
       // Clear the Array and start the request
       IF #wSDOStatus = 12 THEN //Step 12
           FILL_BLK(IN := 0,
                    COUNT := 64,
                    OUT => #bySDODataArray[0]);
           #bSDOReq := TRUE;
           #bSDOWriteDone := FALSE;
           #wSDOStatus := 13; //proceed to Step 13
       END_IF;
       // setup the array data and start WRREC
       IF #wSDOStatus = 13 THEN //Step 13
           #bySDODataArray[0] := 16#f9; //Request Reference
           #bySDODataArray[1] := 16#02; //2 for write PNU
           #bySDODataArray[2] := 16#00; //Axis# is 0 for AKD
           #bySDODataArray[3] := 16#01; // Number of parameters to write at a time
           // Set PNU 916 subindex 5
           #bySDODataArray[4] := 16#10; //Attribute is 0x10
           #bySDODataArray[5] := 16#01; //Number of elements =1
           #bySDODataArray[6] := 16#03; //0x394 for PNU 916
           #bySDODataArray[7] := 16#94; //PNU 916
           #bySDODataArray[8] := 16#00; //subindex
           #bySDODataArray[9] := 16#05; //subindex 5 for 6th word of telegram
           // To PNU 52 (ITIST_GLATT)
           #bySDODataArray[10] := 16#42; //Format =0x42 for Word
           #bySDODataArray[11] := 16#01; //Number of values
           #bySDODataArray[12] := 16#00; //data
           #bySDODataArray[13] := 16#34; //data - Signal #52 (0x34) for ITIST_GLATT (IL.FB)

           #SDOWrite(REQ := #bSDOReq, //do the PNU write
                     ID := #iID,
                     INDEX := 47, //AKD suppors "Record Data 47"
                     LEN := 14,   //data length
                     BUSY => #bSDOWriteBusy,
                     DONE => #bSDOWriteDone,
                     ERROR => #bSDOWriteError,
                     RECORD := #bySDODataArray);
           IF #bSDOWriteBusy THEN
               #bSDOReq := FALSE;
           ELSIF #bSDOWriteDone THEN
               #wSDOStatus := 14; //proceed to Step 14
               //#oInitDone := 1;    //telegram configuration complete
           END_IF;
       END_IF;

       // Set OpMode 
       // Clear the Array and start the request
       IF #wSDOStatus = 14 THEN //Step 14
           FILL_BLK(IN := 0,
                    COUNT := 64,
                    OUT => #bySDODataArray[0]);
           #bSDOReq := TRUE;
           #bSDOWriteDone := FALSE;
           #wSDOStatus := 15; //proceed to Step 15
       END_IF;
       // Set OpMode = 2 Position
       IF #wSDOStatus = 15 THEN //Step 15
           #bySDODataArray[0] := 16#fe; //Request Reference
           #bySDODataArray[1] := 16#02; //2 for write PNU
           #bySDODataArray[2] := 16#00; //Axis# is 0 for AKD
           #bySDODataArray[3] := 16#01; // Number of parameters to write at a time
               // Set PNU 930 subindex 0 (DRV.OPMODE)
           #bySDODataArray[4] := 16#10; //Attribute is 0x10
           #bySDODataArray[5] := 16#01; //Number of elements =1
           #bySDODataArray[6] := 16#03; //0x3A2 for PNU 930 - opmode
           #bySDODataArray[7] := 16#A2; //PNU 930
           #bySDODataArray[8] := 16#00; //subindex 0
           #bySDODataArray[9] := 16#00; //subindex 0
               // To 2 (position mode)
           #bySDODataArray[10] := 16#42; //Format =0x42 for Word
           #bySDODataArray[11] := 16#01; //Number of values
           #bySDODataArray[12] := 16#02; //data
           #bySDODataArray[13] := 16#02; //data - vlaue = 2 for position mode

           #SDOWrite(REQ := #bSDOReq, //do the PNU write
                     ID := #iID,
                     INDEX := 47, //AKD suppors "Record Data 47"
                     LEN := 14,   //data length
                     BUSY => #bSDOWriteBusy,
                     DONE => #bSDOWriteDone,
                     ERROR => #bSDOWriteError,
                     RECORD := #bySDODataArray);
           IF #bSDOWriteBusy THEN
               #bSDOReq := FALSE;
           ELSIF #bSDOWriteDone THEN
               #wSDOStatus := 20; // setup complete - skip to process
               #oInitDone := TRUE;    //telegram configuration complete
           END_IF;
       END_IF;
   END_IF;

   // Read ZSW and set output values
   IF NOT #iInit AND #wSDOStatus > 19 THEN
       #wPNReadStatus := DPRD_DAT(LADDR := #iID,
                                  RECORD => #TG_400.Receive);
       IF #wPNReadStatus = 0 THEN
           #bPNReadError := FALSE;

           #oStatus.%W0 := #TG_400.Receive.ZSW1;
           IF #wSDOStatus > 20 THEN
               #oStatus.%W1 := #wSDOReadValue;
           ELSE
               #oStatus.%W1 := 0;
           END_IF;
           #oPos.%W0 := #TG_400.Receive.XIST_A_1;
           #oPos.%W1 := #TG_400.Receive.XIST_A;
           #oVel := #TG_400.Receive.NIST_A;
           #oCurrent := #TG_400.Receive.ITIST_GLATT;

           #oEnabled := #TG_400.Receive.ZSW1.%X0 AND #TG_400.Receive.ZSW1.%X1 AND #TG_400.Receive.ZSW1.%X2 AND NOT #TG_400.Receive.ZSW1.%X6;
           #oFault := #TG_400.Receive.ZSW1.%X3;
           #oMoving := NOT #TG_400.Receive.ZSW1.%X13 OR #TG_400.Receive.ZSW1.%X14 OR #TG_400.Receive.ZSW1.%X12;
           #oHomed := #TG_400.Receive.ZSW1.%X11;
           IF #TG_400.Send.STW1.%X6 THEN        // Reset the InPos Flag for a minimum of one write cycle
               #oInPos := FALSE;
           ELSE
               #oInPos := #TG_400.Receive.ZSW1.%X10;
           END_IF;
           #oWarning := #TG_400.Receive.ZSW1.%X7;
       ELSE
           #bPNReadError := TRUE;
       END_IF;

   END_IF;

   // Do the write always as the zero Telegramm needs to be send on a init aswell
   #wPNWriteStatus := DPWR_DAT(LADDR := #iID,
                               RECORD := #TG_400.Send);

   // set STW1 and values for the AKD
   IF NOT #iInit AND #wSDOStatus > 19 THEN
       IF #wPNWriteStatus = 0 THEN
           #bPNWriteError := FALSE;

           #TG_400.Send.STW1.%X10 := TRUE;
           IF #TG_400.Receive.ZSW1.%X9 THEN     // PLC has control

               // Do a EStop
               IF #iEStop THEN
                   #TG_400.Send.STW1.%X2 := FALSE;
                   #bEstop := TRUE;
               END_IF;

               // Do a reset
               IF #iReset AND NOT #bResetDone THEN
                   #wSDOStatus := 20;
                   #TG_400.Send.STW1.%X7 := TRUE;
                   #bResetDone := TRUE;
                   #bEstop := FALSE;
                   #wStartReset := #TG_400.Receive.ZSW2;
               END_IF;
               IF ABS(#wStartReset - #TG_400.Receive.ZSW2) > 2 THEN
                   #TG_400.Send.STW1.%X7 := FALSE;
               END_IF;

               // Enable the drive
               IF #iSW_Enable AND NOT #bEstop AND NOT (#bSWEnabled AND #TG_400.Receive.ZSW1.%X6 OR #TG_400.Receive.ZSW1.%X3) THEN
                   IF #TG_400.Receive.ZSW1.%X6 THEN      // Switch on inhibited
                       #TG_400.Send.STW1.%X1 := TRUE;
                       #TG_400.Send.STW1.%X2 := TRUE;
                   ELSE
                       IF #TG_400.Receive.ZSW1.%X0 THEN     // Ready for switiching on
                           #TG_400.Send.STW1.%X0 := TRUE;
                           IF #TG_400.Receive.ZSW1.%X1 THEN       // Switched on
                               #TG_400.Send.STW1.%X3 := TRUE;
                               IF #TG_400.Receive.ZSW1.%X2 THEN       // Operation
                                   #TG_400.Send.STW1.%X12 := TRUE; //turn on real time jogging mode
                                   #bSWEnabled := TRUE;

                                   // Do a Stop
                                   IF #iStop THEN
                                       #TG_400.Send.STW1.%X4 := FALSE;   // Stop active motion task
                                       #TG_400.Send.STW1.%X5 := FALSE;   // Stop active motion task
                                       #TG_400.Send.STW1.%X8 := FALSE;   // Stop jog 1
                                       #TG_400.Send.STW1.%X9 := FALSE;   // Stop jog 2
                                       #TG_400.Send.STW1.%X11 := FALSE;  // Stop homeing
                                       //#TG_400.Send.STW1.%X12 := FALSE;  // Stop real time jogging mode
                                   ELSE

                                       // Do home
                                       IF #iStart_Homing AND NOT #bHomeStarted THEN
                                           #TG_400.Send.HOME_DIST := #iCmdPos.%W1;
                                           #TG_400.Send.HOME_DIST_1 := #iCmdPos.%W0;
                                           #TG_400.Send.STW1.%X11 := TRUE;
                                           #wHomingStartPoint := #TG_400.Receive.ZSW2;
                                           #bHomeStarted := TRUE;
                                       ELSE
                                           IF #TG_400.Receive.ZSW1.%X11 AND #TG_400.Receive.ZSW1.%X13 AND (ABS(#wHomingStartPoint - #TG_400.Receive.ZSW2) > 5) THEN
                                               #TG_400.Send.STW1.%X11 := FALSE;
                                           END_IF;

                                           // Jogging
                                           IF #iStart_Jog AND #iCmdVel <> 0 THEN
                                               #TG_400.Send.STW1.%X8 := TRUE;
                                               //#TG_400.Send.STW1.%X12 := TRUE;

                                               // if the speed input is negative set Bit 13 for reverse direction 
                                               IF #iCmdVel.%X31 = 1 THEN
                                                   #TG_400.Send.STW1.%X13 := TRUE;
                                                   #TG_400.Send.MDI_VELOCITY := (16#ffff - #iCmdVel.%W1 + 1);
                                                   #TG_400.Send.MDI_VELOCITY_1 := (16#ffff - #iCmdVel.%W0 + 1);
                                               ELSE
                                                   #TG_400.Send.STW1.%X13 := FALSE;
                                                   #TG_400.Send.MDI_VELOCITY := #iCmdVel.%W1;
                                                   #TG_400.Send.MDI_VELOCITY_1 := #iCmdVel.%W0;
                                               END_IF;

                                               #TG_400.Send.MDI_ACC := #iCmdAcc;
                                               #TG_400.Send.MDI_DEC := #iCmdDec;
                                           ELSE
                                               #TG_400.Send.STW1.%X8 := FALSE;
                                               //#TG_400.Send.STW1.%X12 := FALSE;

                                               // Interrupt a move
                                               IF #iMT_Pause THEN
                                                   #TG_400.Send.STW1.%X5 := FALSE;    // intermediate stop, motion is paused and will continue when the pause is lifted
                                               ELSE
                                                   #TG_400.Send.STW1.%X5 := TRUE;    // No intermediate stop
                                               END_IF;

                                               // Reset the rising edge of the start bit to be read for the next task
                                               IF #TG_400.Receive.ZSW1.%X12 OR ABS(#wStartMove - #TG_400.Receive.ZSW2) > 62 THEN //if start command has been acknowledged, or >62 telegram transmissions
                                                   #bStartMoveDone := TRUE; // the process to start the move has been completed
                                                   #TG_400.Send.STW1.%X6 := FALSE; //turn off the start bit
                                               END_IF;
                                               // Move
                                               IF #iStart_Move AND NOT #bStartMove THEN
                                                   #TG_400.Send.MDI_MOD := #iMT_MoveType;   // 1 = absolute, 0 = relative
                                                   #TG_400.Send.SATZANW := #iMTNum;      // 0x8000 = direct motion task, otherwise select a motion task from the AKD
                                                   #TG_400.Send.MDI_TARPOS := #iCmdPos.%W1;
                                                   #TG_400.Send.MDI_TARPOS_1 := #iCmdPos.%W0;
                                                   #TG_400.Send.MDI_VELOCITY := #iCmdVel.%W1;
                                                   #TG_400.Send.MDI_VELOCITY_1 := #iCmdVel.%W0;
                                                   #TG_400.Send.MDI_ACC := #iCmdAcc;
                                                   #TG_400.Send.MDI_DEC := #iCmdDec;
                                                   #TG_400.Send.STW1.%X4 := TRUE;    // Do not reject traversing task
                                                   #TG_400.Send.STW1.%X5 := TRUE;    // No intermediate stop
                                                   #TG_400.Send.STW1.%X6 := TRUE;    // Start the move

                                                   #bStartMove := TRUE; // the process to start the move has been started but not completed
                                                   #bStartMoveDone := FALSE; // the process to start the move has not been completed
                                                   #wStartMove := #TG_400.Receive.ZSW2;
                                               END_IF; //If Start move

                                           END_IF; //If Start Jog
                                       END_IF; //If Start Homing
                                   END_IF; // If Stop
                               END_IF; // If ZSW1 bit2 Operation Enabled
                           END_IF; // If ZSW1 bit1 Switched On
                       END_IF; // If ZSW1 bit0 Ready for Switch On
                   END_IF; // If ZSW1 bit6 Switch-On Inhibited

                   // If the axis gets disabled all the corresponding motion signals have to be reset    
               ELSE
                   #bSWEnabled := FALSE;

                   #TG_400.Send.STW1.%X0 := FALSE;
                   #TG_400.Send.STW1.%X1 := FALSE;
                   #TG_400.Send.STW1.%X2 := FALSE;
                   #TG_400.Send.STW1.%X3 := FALSE;
                   #TG_400.Send.STW1.%X4 := FALSE;
                   #TG_400.Send.STW1.%X5 := FALSE;
                   #TG_400.Send.STW1.%X6 := FALSE;
                   #TG_400.Send.STW1.%X8 := FALSE;
                   #TG_400.Send.STW1.%X9 := FALSE;
                   #TG_400.Send.STW1.%X11 := FALSE;
                   #TG_400.Send.STW1.%X12 := FALSE;
               END_IF; //If Enable
           END_IF; // ZSW1 bit9 PLC has control
       ELSE
           #bPNWriteError := TRUE;
       END_IF; //If #wPNWriteStatus = 0

       // Read drive faults and warning on occurens
       IF #oFault THEN
           // If alarm is not read yet: start read
           IF NOT #wSDOStatus.%X6 AND NOT #bSDOStatusReadActive THEN
               #wSDOStatus := 64;
               #wSDOAddress := 16#09AD;     // Read PNU 2477 (DRV.FAULT1)
               #bSDOStatusReadActive := TRUE;
           END_IF;

           // If warning is not read yet: start read
       ELSIF #oWarning THEN
           IF NOT #wSDOStatus.%X5 AND NOT #bSDOStatusReadActive THEN
               #wSDOStatus := 32;
               #wSDOAddress := 16#0AE7;    // Read PNU2791 (DRV.WARNING1)
               #bSDOStatusReadActive := TRUE;
           END_IF;
       ELSE
           IF NOT #bSDOStatusReadActive THEN
               #wSDOStatus := 20;
           END_IF;
       END_IF; //IF #oFault

       // start the reading signal
       IF #wSDOStatus >= 32 THEN
           // Always clean out old values first
           IF #bSDOWriteBusy THEN
               #bSDOReq := FALSE;
           ELSE
               FILL_BLK(IN := 0,
                        COUNT := 64,
                        OUT => #bySDODataArray[0]);
               #bSDOReq := TRUE;
               #bSDOWriteDone := FALSE;
           END_IF;
           // Start the read cylce to the corrsponding PNU 
           IF #wSDOStatus = 32 OR #wSDOStatus = 64 THEN
               #bySDODataArray[0] := #wSDOStatus.%B0;
               #bySDODataArray[1] := 16#01;
               #bySDODataArray[2] := 16#00;
               #bySDODataArray[3] := 16#01;

               #bySDODataArray[4] := 16#10;
               #bySDODataArray[5] := 16#01;
               #bySDODataArray[6] := #wSDOAddress.%B1;
               #bySDODataArray[7] := #wSDOAddress.%B0;
               #bySDODataArray[8] := 16#00;
               #bySDODataArray[9] := 16#00;

               #SDOWrite(REQ := #bSDOReq,
                         ID := #iID,
                         INDEX := 47,
                         LEN := 14,
                         BUSY => #bSDOWriteBusy,
                         DONE => #bSDOWriteDone,
                         ERROR => #bSDOWriteError,
                         RECORD := #bySDODataArray);
               IF #bSDOWriteDone THEN
                   #wSDOStatus := #wSDOStatus + 1;
               END_IF;
           END_IF; //IF #wSDOStatus = 32 OR #wSDOStatus = 64

           // read the value back
           IF #wSDOStatus = 33 OR #wSDOStatus = 65 THEN
               #SDORead(REQ := #bSDOReq,
                        ID := #iID,
                        INDEX := 47,
                        MLEN := 14,
                        BUSY => #bSDOReadBusy,
                        VALID => #bSDOReadDone,
                        ERROR => #bSDOReadError,
                        RECORD := #bySDODataArray);
               IF #bSDOReadDone THEN
                   IF #bySDODataArray[4] = 66 THEN               // if the read signal is a Word use Byte 6&7
                       #wSDOReadValue.%B0 := #bySDODataArray[7];
                       #wSDOReadValue.%B1 := #bySDODataArray[6];
                   ELSE                                        // if the read signal is a DWord use Byte 8&9
                       #wSDOReadValue.%B0 := #bySDODataArray[9];
                       #wSDOReadValue.%B1 := #bySDODataArray[8];
                   END_IF;
                   IF #wSDOReadValue = 0 THEN  // If the read value is zero repeat the read cycle
                       #wSDOStatus := #wSDOStatus - 1;
                   ELSE
                       #wSDOStatus := #wSDOStatus + 1;
                       #bSDOStatusReadActive := FALSE;
                   END_IF;
               END_IF; //IF #bSDOReadDone
           END_IF; //IF #wSDOStatus = 33 OR #wSDOStatus = 65
       END_IF; //IF #wSDOStatus >= 32
   END_IF; //IF NOT #iInit AND #wSDOStatus > 19

   //  check for rising edge for the input parameters
   IF NOT #iReset AND #bResetDone THEN
       #bResetDone := FALSE;
   END_IF;
   IF NOT #iStart_Homing AND #bHomeStarted THEN
       #bHomeStarted := FALSE;
   END_IF;
   IF NOT #iStart_Move AND #bStartMove AND #bStartMoveDone AND NOT #TG_400.Receive.ZSW1.%X12 THEN
       #bStartMove := FALSE;
       #bStartMoveDone := FALSE;
   END_IF;

   // fault detection/handling within the bloc
   IF #bPNReadError OR #bPNWriteError OR #bSDOReadError OR #bSDOWriteError THEN
       #oError := TRUE;
       IF #bPNReadError THEN
           #oStatus := #wPNReadStatus; //indicates internal FB error
       END_IF;
       IF #bPNWriteError THEN
           #oStatus := #wPNWriteStatus; //indicates internal FB error
       END_IF;
   ELSIF #wSDOStatus > 19 THEN
       #oError := FALSE;
   END_IF;
END_FUNCTION_BLOCK

// folder: AKD/PNU

FUNCTION_BLOCK "AKD_PNU_v02"   // FB15, SCL
TITLE = AKD_PNU_v02
{ S7_Optimized_Access := 'FALSE' }
AUTHOR : jcoleman
FAMILY : PNU
VERSION : 2.0
// This function block uses the Parameter Access channel to read and write PNU parameters values.
   VAR_INPUT
      iID : Hw_Io;   // unique connection ID
      iStartRequest : Bool;   // start Read or Write
      iRequestType : Bool;   // 0 = Read; 1 = Write
      iFormat : Int;   // Datatype 0x41 = Byte, 0x42 = Word, 0x43 = DWord
      iPNUnumber : Word;   // PNU address
      iPNUsubIndex : Word;   // PNU Subindex
   END_VAR
   VAR_OUTPUT
      oActive : Bool;   // request in progress
      oDone : Bool;   // request finished
      oError : Bool;   // request failed
      oStatus : DWord;   // status of the failed function
   END_VAR
   VAR_IN_OUT
      ioData : DWord;
   END_VAR
   VAR
      PNURead : RDREC;
      PNUWrite : WRREC;
      bDoWrite : Bool;
      bDoRead : Bool;
      byReadArray : Array[0..147] of Byte;
      byWriteArray : Array[0..31] of Byte;
      bPNUWriteBusy : Bool;
      bPNUWriteDone : Bool;
      bPNUWriteError : Bool;
      dwPNUWriteStatus : DWord;
      bPNUReadBusy : Bool;
      bPNUReadDone : Bool;
      bPNUReadError : Bool;
      dwPNUReadStatus : DWord;
      wDataLenght : Word;
      bReqActive : Bool;
      wLenght : Word;
      byReference : Byte;
      bReadActive : Bool;
      bWriteActive : Bool;
   END_VAR
BEGIN
   ////////////////////////////////////////////////////////////////////////////////////////////////////////
   // Communication module between a Kollmorgen AKD and S7-1200/1500 PLC, for direct parameter access
   // 
   // Version  When        Who         What
   // ---------------------------------------------
   // V 2.000  17.07.06    JColeman KM Changed input and output names
   // V 1.000  17.09.15    MRupf KM    Conversion to TIA V13 SP1
   // V 0.005  14.07.15    MRupf KM    Automatic format check for read values
   // V 0.004  06.07.15    MRupf KM    oDone and oActive Trigger corrected
   // V 0.002  26.02.15    MRupf KM    iSubIndex added
   // V 0.001  18.02.15    MRupf KM    first version
   //////////////////////////////////////////////////////////////////////////////////////////////////////////

   // Set the output in error case and only reset with new req
   IF #bPNUReadError OR #bPNUWriteError OR (#iFormat - 16#41 < 0) OR (#iFormat - 16#43 > 0) THEN
       #oError := TRUE;
       IF #bPNUReadError THEN
           #bDoRead := FALSE;
           #oStatus := #dwPNUReadStatus;
       END_IF;
       IF #bPNUWriteError THEN
           #bDoWrite := FALSE;
           #oStatus := #dwPNUWriteStatus;
       END_IF;
   END_IF;

   // Request edge starts a new call if none active
   IF #iStartRequest AND NOT #bReqActive THEN
       #byReference := #byReference + 1;     // Every request gets a new reference for debuging purpose
       IF #byReference = 0 THEN
           #byReference := #byReference + 1;
       END_IF;

       // Reset all the status bit with every request
       #oActive := TRUE;
       #oDone := FALSE;
       #oError := FALSE;
       #oStatus := 0;

       FILL_BLK(IN := 0,
                COUNT := 16,
                OUT => #byWriteArray[0]);

       FILL_BLK(IN := 0,
                COUNT := 148,
                OUT => #byReadArray[0]);

       // Set the data to start a PNU write request
       IF #iRequestType THEN
           #byWriteArray[0] := #byReference;      // Byte 0        reference
           #byWriteArray[1] := 16#02;            // Byte 1        Request ID (2 = write) 
           #byWriteArray[2] := 16#00;            // Byte 2        Axis (0)
           #byWriteArray[3] := 16#01;            // Byte 3        Number of parameters
           #byWriteArray[4] := 16#10;            // Byte 4        Attribute
           #byWriteArray[5] := 16#01;            // Byte 5        Number of elements
           #byWriteArray[6] := #iPNUnumber.%B1;        // Byte 6&7      PNU number
           #byWriteArray[7] := #iPNUnumber.%B0;        // Byte 6&7      PNU number
           #byWriteArray[8] := #iPNUsubIndex.%B1;    // Byte 8&9      Subindex (0)
           #byWriteArray[9] := #iPNUsubIndex.%B0;    // Byte 8&9      Subindex (0)
           #byWriteArray[10] := #iFormat;         // Byte 10       Format
           #byWriteArray[11] := 16#01;           // Byte 11       Number of values

           // Set the lenght automatically according to the Format
           IF #iFormat = 16#41 THEN
               #wLenght := 16#0E;
               #byWriteArray[12] := #ioData.%B0;    // Byte 12    Value
           ELSE
               IF #iFormat = 16#42 THEN
                   #wLenght := 16#10;
                   #byWriteArray[12] := #ioData.%B1;    // Byte 12&13    Value
                   #byWriteArray[13] := #ioData.%B0;    // Byte 12&13    Value
               ELSE
                   IF #iFormat = 16#43 THEN
                       #wLenght := 16#14;
                       #byWriteArray[12] := #ioData.%B3;    // Byte 12&13    Value
                       #byWriteArray[13] := #ioData.%B2;    // Byte 12&13    Value
                       #byWriteArray[14] := #ioData.%B1;    // Byte 14&15    Value
                       #byWriteArray[15] := #ioData.%B0;    // Byte 14&15    Value
                   END_IF;
               END_IF;
           END_IF;

           #bDoWrite := TRUE;

       // Set the data to start a PNU read request 
       ELSE
           #byWriteArray[0] := #byReference;      // Byte 0       reference
           #byWriteArray[1] := 16#01;            // Byte 1       Request ID (1 = read)
           #byWriteArray[2] := 16#00;            // Byte 2       Axis (0)
           #byWriteArray[3] := 16#01;            // Byte 3       Number of parameters
           #byWriteArray[4] := 16#10;            // Byte 4       Attribute
           #byWriteArray[5] := 16#01;            // Byte 5       Number of elements
           #byWriteArray[6] := #iPNUnumber.%B1;        // Byte 6&7     PNU number
           #byWriteArray[7] := #iPNUnumber.%B0;        // Byte 6&7     PNU number
           #byWriteArray[8] := #iPNUsubIndex.%B1;    // Byte 8&9     Subindex (0)
           #byWriteArray[9] := #iPNUsubIndex.%B0;    // Byte 8&9     Subindex (0)

           #ioData := 0;
           #bDoWrite := TRUE;
       END_IF;

     #bReqActive := TRUE;
   END_IF;

   // Start the request
   #PNUWrite(REQ := #bDoWrite,
             ID := #iID,
             INDEX := 47,
             LEN := #wLenght,
             BUSY => #bPNUWriteBusy,
             DONE => #bPNUWriteDone,
             ERROR => #bPNUWriteError,
             STATUS => #dwPNUWriteStatus,
             RECORD := #byWriteArray);

   // Read the answer 
   #PNURead(REQ := #bDoRead,
            ID := #iID,
            INDEX := 47,
            MLEN := 148,
            BUSY => #bPNUReadBusy,
            VALID => #bPNUReadDone,
            ERROR => #bPNUReadError,
            STATUS => #dwPNUReadStatus,
            LEN => #wDataLenght,
            RECORD := #byReadArray);

   // Copie the read data to the output
   IF NOT #iRequestType THEN
       // Set the data automatically according to the Format
       IF #byReadArray[4] = 16#41 THEN
           #ioData.%B0 := #byReadArray[6];    // Byte 10    Value
           #ioData.%B1 := 0;
           #ioData.%B2 := 0;
           #ioData.%B3 := 0;
       ELSE
           IF #byReadArray[4] = 16#42 THEN
               #ioData.%B0 := #byReadArray[7];    // Byte 12&13    Value
               #ioData.%B1 := #byReadArray[6];    // Byte 12&13    Value
               #ioData.%B2 := 0;
               #ioData.%B3 := 0;
           ELSE
               IF #byReadArray[4] = 16#43 THEN
                   #ioData.%B0 := #byReadArray[9];    // Byte 12&13    Value
                   #ioData.%B1 := #byReadArray[8];    // Byte 12&13    Value
                   #ioData.%B2 := #byReadArray[7];    // Byte 14&15    Value
                   #ioData.%B3 := #byReadArray[6];    // Byte 14&15    Value
               END_IF;
           END_IF;
       END_IF;
   END_IF;

   // Reset the request bit for the read and write
   IF #bPNUWriteBusy THEN
       #bDoWrite := FALSE;
       #bWriteActive := TRUE;
   ELSIF #bPNUWriteDone THEN
       #bDoRead := TRUE;
       #bWriteActive := FALSE;
   END_IF;
   IF #bPNUReadBusy THEN
       #bDoRead := FALSE;
       #bReadActive := TRUE;
   ELSIF #bPNUReadDone THEN
       #bReadActive := FALSE;
   END_IF;

   // Set the output bit after a request is processed
   IF #oActive AND #byReadArray[0] = #byReference THEN
       #oActive := FALSE;
       #oDone := TRUE;
   END_IF;

   // Check for the rising edge of req
   IF NOT #iStartRequest AND #bReqActive THEN
       #bReqActive := FALSE;
   END_IF;
END_FUNCTION_BLOCK

// folder: MQTT

FUNCTION_BLOCK "LMqtt_Publisher_1"   // FB8, SCL
{ S7_Optimized_Access := 'TRUE' }
VERSION : 0.1
   VAR_INPUT
      enable : Bool;
      publish : Bool;
      tcpConnParam : "typeTcpConnParam";
      mqttParam : "typeMqttParam_1";
   END_VAR
   VAR_OUTPUT
      tcpEstablished : Bool;
      mqttEstablished : Bool;
      published : Bool;
      busy : Bool;
      error : Bool;
      status : DWord;
      statusID : Int;
   END_VAR
   VAR
      statTcpConnParam : TCON_IP_v4;
      instTcpConnect : TCON;
      instTcpSend : TSEND;
      instTcpRCV : TRCV;
      instTcpDisconnect : TDISCON;
      instWatchDog : TON_TIME;
      instKeepAlive : TON_TIME;
      statStateMQTT : Int;
      statStateMQTTinternal : Int;
      statStateTCP : Int;
      statLastState : Int;
      statConnectLenght : Int;
      statCorrectOffset : Int;
      statSendLenght : Int;
      statConnectEncodedLenght : Int;
      statConnectLenghtOffset : Int;
      statKeepAliveTime : Time;
      statI : Int;
      statPacketID : Word;
      statPacketIDAck : Word;
      statRcvLen : UDInt;
      statPublishOld : Bool;
      statReConnect : Bool;
      statEnableOld : Bool;
      statMqttResetOld : Bool;
      statTriggerWatchDog : Bool;
      statTriggerKeepAlive : Bool;
      statNewDataRcv : Bool;
      statKeepAliveOff : Bool;
      statSendBuffer : Array[1..1000] of Byte;
      statRcvBuffer : Array[1..200] of Byte;
   END_VAR
   VAR_TEMP
      tempStringToChar : Array[0..2000] of Char;
      tempCountChars : UInt;
      tempLenght : Word;
      test : Array[0..1] of Int;
      testarray : Array[0..1] of WChar;
   END_VAR
   VAR CONSTANT
      TCP_PARAM : Int := 1;
      TCP_DISCONNECT : Int := -1;
      TCP_ERROR : Int := -2;
      TCP_CONNECTED : Int := 3;
      TCP_CONNECTING : Int := 2;
      MQTT_CONNECT_FLAG_CHECK : Int := 10;
      MQTT_CONNECT : Int := 11;
      MQTT_PUBLISH : Int := 13;
      MQTT_DISCONNECT : Int := 15;
      MQTT_CONNACK : Int := 12;
      MQTT_PUBACK : Int := 14;
      MQTT_PING : Int := 17;
      MQTT_PINGRESP : Int := 18;
      MQTT_PUBREL : Int := 19;
      MQTT_PUBCOMP : Int := 20;
      MQTT_IDLE : Int;
      MQTT_CONNECTED : Int := 16;
      MQTT_DISCONNECTED : Int := -11;
      MQTT_ERROR : Int := -12;
      IDLE : Int;
      TIME_MONITORING : Int := 20;
      WATCHDOG_TIME : Time := t#30s;
      MQTT_MSG_TYPE_CONNACK : Int := 32;
      MQTT_MSG_TYPE_DISCONNECT : Int := 224;
      MQTT_MSG_TYPE_PUBACK : Int := 64;
      MQTT_MSG_TYPE_PUBREC : Int := 80;
      MQTT_MSG_TYPE_PUBCOM : Int := 112;
      MQTT_MSG_TYPE_PING : Int := 192;
      MQTT_MSG_TYPE_PINGRESP : Int := 208;
      MQTT_CONNACK_ACCEPTED : Int;
      MQTT_PORT : Word := 16#22B3;
      MQTT_PROTOCOL_NAME : String := 'MQTT';
      MQTT_ERROR_WILL_FLAG : Word := 16#80F0;
      MQTT_ERROR_QOS_FLAG : Word := 16#80F1;
      MQTT_ERROR_PACKETID : Word := 16#80F2;
      MQTT_ERROR_KEEPALIVE : Word := 16#80F3;
   END_VAR
   // statTcpConnParam.ActiveEstablished := true;
BEGIN
   //=============================================================================
   //SIEMENES AG
   //(c)Copyright 2016 All Rights Reserved
   //-----------------------------------------------------------------------------
   //Library:       (that the source is dedicated to)
   //Tested with:   (target system with FW Version)
   //Engineering:   TIA Portal V15
   //Restrictions:  (OB types, etc.)
   //Requirements:  (hardware, technological package, memory needed, etc.)
   //Functionality: MQTT
   //-----------------------------------------------------------------------------
   //Change log table:
   //Version  Date       Expert in charge Changes applied
   //01.00.00 dd.mm.yyyy (name of expert) First released version
   //=============================================================================
   //Establish TCP Connection to be ready for MQTT

   IF #enable
       AND NOT #statEnableOld
   THEN
       #statStateTCP := #TCP_PARAM;
       #statStateMQTT := #MQTT_DISCONNECTED;
       #instWatchDog.IN := false;
       #statPublishOld := #publish;
       #error := 0;
       #status := 0;
       #statusID := 0;
   END_IF;

   IF NOT #enable
       AND #statEnableOld
   THEN
       IF #statStateTCP = #TCP_CONNECTED AND
           #statStateMQTT = #MQTT_DISCONNECTED
       THEN
           #statStateTCP := #TCP_DISCONNECT;
       END_IF;
       IF #statStateTCP = #TCP_CONNECTED AND
           #statStateMQTT <> #MQTT_DISCONNECTED
       THEN
           #statStateMQTT := #MQTT_DISCONNECT;
       END_IF;
       IF #statStateTCP = #TCP_CONNECTING
           OR  #statStateTCP = #IDLE
       THEN

           #statStateMQTT := #MQTT_DISCONNECTED;
           #statStateTCP := #IDLE;
       END_IF;
   END_IF;

    #instWatchDog(IN := #statTriggerWatchDog,PT := #WATCHDOG_TIME);

   REGION State maschine TCP
       CASE #statStateTCP OF
           #IDLE:
               IF NOT #error
               THEN
                   #status := 0;
                   #statusID := 0;

               END_IF;
               #statTcpConnParam.ID := #tcpConnParam.connectionID;
               #instTcpDisconnect(ID := #statTcpConnParam.ID);
               #instTcpConnect(ID := #statTcpConnParam.ID,
                               CONNECT := #statTcpConnParam);
               #published := 0;
               #busy := false;
               #mqttEstablished := false;
               #statMqttResetOld := 0;
               #tcpEstablished := false;
               #statStateMQTT := #MQTT_DISCONNECTED;
               #statStateMQTTinternal := #IDLE;
               #statTriggerWatchDog := false;
               #statTriggerKeepAlive := 0;
               IF #statLastState=#TCP_DISCONNECT
               THEN
                   #error := 0;
                   END_IF;
           #TCP_CONNECTED:
               ;
               //Check TCP Connection
               IF #instTcpRCV.STATUS > w#16#80C0
               THEN
                   #statStateTCP := #TCP_ERROR;
                   #statusID := #TCP_CONNECTED;
               END_IF;
               #statLastState := #TCP_CONNECTED;
           #TCP_PARAM:
               #statTcpConnParam.InterfaceId := #tcpConnParam.hwIdentifier;
               #statTcpConnParam.ID := #tcpConnParam.connectionID;
               #statTcpConnParam.LocalPort := #tcpConnParam.localPort;
               #statTcpConnParam.RemotePort := #tcpConnParam.mqttPort;
               #statTcpConnParam.ActiveEstablished := true;
               #statTcpConnParam.RemoteAddress.ADDR[1] := #tcpConnParam.ipAdressBroker[0];
               #statTcpConnParam.RemoteAddress.ADDR[2] := #tcpConnParam.ipAdressBroker[1];
               #statTcpConnParam.RemoteAddress.ADDR[3] := #tcpConnParam.ipAdressBroker[2];
               #statTcpConnParam.RemoteAddress.ADDR[4] := #tcpConnParam.ipAdressBroker[3];

             #statStateTCP := #TCP_CONNECTING;
           #TCP_CONNECTING:
               REGION TCP Connect
                   #statTriggerWatchDog := true;
                   #instTcpConnect.REQ := NOT #instTcpConnect.REQ XOR #instTcpConnect.BUSY;
                   #instTcpConnect(ID := #statTcpConnParam.ID,
                                   CONNECT := #statTcpConnParam);

                   IF (#instTcpConnect.DONE)
                       AND (#instTcpConnect.BUSY = 0)
                       AND (#instTcpConnect.REQ)
                   THEN
                       #instTcpConnect.REQ := false;
                       #tcpEstablished := true;
                       #statStateTCP := #TCP_CONNECTED;
                       #statTriggerWatchDog := false;
                   ELSIF (#instTcpConnect.ERROR)
                   THEN
                       #statusID := #TCP_CONNECTING;
                       #instTcpConnect.REQ := false;
                       #statStateTCP := #TCP_ERROR;
                   END_IF;
               END_REGION

           #TCP_DISCONNECT:
               REGION TCP Disconnect
                   #instTcpDisconnect.REQ := NOT #instTcpDisconnect.REQ XOR #instTcpDisconnect.BUSY;
                   #statTriggerWatchDog := false;
                   #instTcpDisconnect(ID := #statTcpConnParam.ID);

                   IF (#instTcpDisconnect.DONE)
                   THEN
                       //Done with success
                       #instTcpDisconnect.REQ := false;
                       #statLastState := #TCP_DISCONNECT;
                       #statStateTCP := #IDLE;
                   ELSIF (#instTcpDisconnect.ERROR)
                   THEN
                       #statusID := #TCP_DISCONNECT;
                       #instTcpDisconnect.REQ := false;
                       #statStateTCP := #TCP_ERROR;
                   END_IF;
               END_REGION
               ;
           #TCP_ERROR:
               REGION Errorhandling
                   #error := true;
                   #statStateMQTT := #MQTT_DISCONNECTED;
                   #statStateMQTTinternal := #IDLE;
                   #tcpEstablished := false;
                   #mqttEstablished := false;
                   #published := false;
                   #statTriggerWatchDog := false;
                   #instTcpConnect.REQ := false;
                       CASE #statusID OF
                           #TCP_CONNECTING:
                               #statStateTCP := #IDLE;
                               #status := #instTcpConnect.STATUS;
                           #TCP_CONNECTED:
                               #statStateTCP := #TCP_DISCONNECT;
                               #status := #instTcpRCV.STATUS;
                           #TCP_DISCONNECT:
                               //pointless for a retry at TDISCON
                               #statStateTCP := #IDLE;
                               #status := #instTcpDisconnect.STATUS;
                           #TIME_MONITORING:
                               IF (#statLastState = #TCP_CONNECTED)
                               THEN
                                   #statStateTCP := #TCP_DISCONNECT;
                                   #status := #instTcpRCV.STATUS;
                               ELSE
                                   #statStateTCP := #IDLE;
                                   #status := #instTcpConnect.STATUS;
                               END_IF;
                           ELSE
                               ;
                       END_CASE;
               END_REGION
               ;
           ELSE
               ;
       END_CASE;
   END_REGION
   #statEnableOld := #enable;
   REGION WatchDog
       IF #instWatchDog.Q = true
       THEN
           #statStateTCP := #TCP_ERROR;
           #statusID := #TIME_MONITORING;
       END_IF;
   END_REGION

   REGION OUC blocks

       #instTcpSend(ID:=#statTcpConnParam.ID,
                     DATA:=#statSendBuffer);
        #instTcpRCV(EN_R:=true,
                    ID:=#statTcpConnParam.ID,
                   LEN:=0,
                   ADHOC:=1,
                   RCVD_LEN=>#statRcvLen,
                   DATA:=#statRcvBuffer);
       IF #instTcpRCV.RCVD_LEN > 0 THEN
           #statNewDataRcv := 1;
       END_IF;

   END_REGION

   //Bring Statemachine in a definded state, if TCP Connection breaks
   IF #statStateMQTT > 0 AND
       #statStateTCP <> #TCP_CONNECTED
   THEN
       #statStateMQTT := #MQTT_DISCONNECTED;
       #instTcpSend.REQ := 0;
   END_IF;

   //MQTT makes no sense without an established TCP
   IF NOT (#statStateTCP = #TCP_CONNECTED)
   THEN
       RETURN;
   END_IF;




    #instKeepAlive(IN := #statTriggerKeepAlive,
                   PT := #statKeepAliveTime);
       CASE #statStateMQTT OF
           #MQTT_DISCONNECTED:
               #mqttEstablished := false;
               #statPublishOld := #publish;
               #statStateMQTT := #MQTT_CONNECT_FLAG_CHECK;
               #statStateMQTTinternal := #IDLE;
               #statTriggerKeepAlive := 0;
               #statKeepAliveOff := false;
               #statPacketID := #mqttParam.packetIdentifier;

           #MQTT_CONNECT_FLAG_CHECK:
               #busy := 1;
               //validate flags
               IF #mqttParam.connectFlag.willRetain
                   AND NOT #mqttParam.connectFlag.will
               THEN
                   #statStateMQTT := #MQTT_ERROR;
                   #statusID := #MQTT_CONNECT_FLAG_CHECK;
                   #status := #MQTT_ERROR_WILL_FLAG;
               ELSE
                   IF NOT #mqttParam.connectFlag.will
                       AND (#mqttParam.connectFlag.willQoS_1 OR #mqttParam.connectFlag.willQoS_2)
                   THEN
                       #statStateMQTT := #MQTT_ERROR;
                       #statusID := #MQTT_CONNECT_FLAG_CHECK;
                       #status := #MQTT_ERROR_QOS_FLAG;
                   ELSE
                       IF (#mqttParam.connectFlag.willQoS_1
                           AND #mqttParam.connectFlag.willQoS_2)
                       THEN
                           #statStateMQTT := #MQTT_ERROR;
                           #statusID := #MQTT_CONNECT_FLAG_CHECK;
                           #status := #MQTT_ERROR_QOS_FLAG;
                       ELSE;
                        #statStateMQTT := #MQTT_CONNECT;
                       END_IF;
                   END_IF;

